// TIA Portal project "g" (V14) (continued)

       REGION Collect-statistics
           // Operating time cnt. (#t_diff will always be zero, if the feature is disabled)
           #devices[#c].operation_time += SEL(G := #devices[#c].in_operation
                                              AND #conf.enable_operation_time_cnt,
                                              IN0 := 0, IN1 := USINT_TO_UDINT(#t_diff));
           // Count number of devices in operation.
           #info.devices_in_operation += BOOL_TO_UINT(#devices[#c].in_operation);
           // Count number of devices in standby.
           #info.devices_standby +=
           BOOL_TO_UINT(#devices[#c].available
                        AND NOT #devices[#c].Q); // NOT #devices[#c].in.in_operation
           // Count number of devices started.
           #info.devices_started += BOOL_TO_UINT(#devices[#c].Q);
       END_REGION
   END_FOR;

   // Some info (for hmi)
   #settings.info.total := DINT_TO_UINT(#upper - #lower + 1);

   // If for some reason, the number operating devies can be limited to less
   // then available
   #settings.max_devices_same_time := // A setting.
   LIMIT(MN := 1,
         IN := #settings.max_devices_same_time,
         MX := #settings.info.total);

   // Force min value for param.
   #settings.max_diff_operating.sec :=
   MAX(IN1 := 60, IN2 := #settings.max_diff_operating.sec);

   // Timers for adding and removing devices for operation.

   #timer_stop.TON(IN := #input < #settings.stop.limit AND NOT #reset_timers,
                   PT := #settings.stop.delay,
                   Q => #timer_stop_q);
   #timer_start.TON(IN := #input > #settings.start.limit AND NOT #reset_timers,
                    PT := #settings.start.delay,
                    Q => #timer_start_q);

   REGION start-stopp
       // Stoping a device
       IF NOT #settings.bypass // The bypass-function turn on all outputs. 
           AND #candidates.stop.index <> #NO_CANDIDATE // A device is available 
           AND (#info.devices_in_operation > 1 // Can't remove last device in operation
           (* *)OR NOT #conf.at_least_one)  // Possible to disable the feature
           AND (
           (* *)#info.devices_in_operation > #settings.max_devices_same_time
           (* *)OR #timer_stop_q // If #input below a certain value for a certain time
           (* *)OR #settings.stop.force  // Used to stop the next device (hmi)
           (* *)OR #boost_start < 0)
       THEN
           #devices[#candidates.stop.index].Q := false; // Disable one device
           RESET_TIMER(#timer_stop);
           #oper := -1;
           // Increase var until zero.
           #boost_start := SEL(G := #boost_start < 0, IN0 := 0, IN1 := #boost_start + 1);

           // Start a devices.
       ELSIF #candidates.start.index <> #NO_CANDIDATE // A device is available 
           AND #info.devices_in_operation < #settings.max_devices_same_time
           AND #input > 0 AND (
           (* *)#info.devices_in_operation < 1 // At least one device operating
           (*      *)AND #conf.at_least_one // Possible to disable the feature
           (* *)OR #timer_start_q // If #input above a certain value for a certain time
           (* *)OR #settings.start.force // Used to starp the next device (hmi)
           (* *)OR #boost_start > 0)
       THEN
           #devices[#candidates.start.index].Q := true; // Enable one more device
           RESET_TIMER(#timer_start);
           #oper := 1;
           // Decrease var until zero.
           #boost_start := SEL(G := #boost_start > 0, IN0 := 0, IN1 := #boost_start - 1);

           // Change operating device, if the operating-time between two devies is to large.
       ELSIF #settings.max_diff_operating.enable
           AND #candidates.start.index <> #NO_CANDIDATE // A candidate is available to be started
           AND #candidates.stop.index <> #NO_CANDIDATE // A candidate is available to be stoped
           AND (#candidates.stop.operation_time - #candidates.start.operation_time >
           (* *)#settings.max_diff_operating.sec) // And the difference is to large.
       THEN
           // Stop the device with most operating time and start the devices with
           // least operating time.
           #devices[#candidates.stop.index].Q := false;
           #devices[#candidates.start.index].Q := true;
       END_IF;
   END_REGION

   // Update vars, after start or stop a device. (above)
   #info.devices_in_operation += SINT_TO_UINT(#oper);
   #info.devices_started += SINT_TO_UINT(#oper);
   #info.devices_standby -= SINT_TO_UINT(#oper);

   // Transfer values to hmi-vars
   #settings.info.in_operation := #info.devices_in_operation;
   #settings.info.started := #info.devices_started;
   #settings.info.standby := #info.devices_standby;

   #settings.info.input := #input;

   // Information has been recived, so now back to default values.
   #set := -1;
   #settings.start.force := false;
   #settings.stop.force := false;
   #settings.boostStart.reset := false;

   // https://github.com/rexhip/
END_FUNCTION_BLOCK

// folder: Library/Alternating/Load balancer/Blocks and UDT's/Internal

FUNCTION "boost_start" : Void   // FC25, SCL
{ S7_Optimized_Access := 'TRUE' }
VERSION : 0.1
   VAR_INPUT
      t_diff : USInt;
      start : Bool;
   END_VAR
   VAR_OUTPUT
      reset_timers : Bool;
   END_VAR
   VAR_IN_OUT
      devices : Array[*] of "load_balancer_device_udt";
      settings : "load_balancer_settings_udt";
      info : "load_balancer_info_udt";
      boost_start : SInt;
      set : SInt;
   END_VAR
   VAR_TEMP
      c : DInt;
      u : DInt;
      lower : DInt;
   END_VAR
BEGIN
   #lower := LOWER_BOUND(ARR := #devices, DIM := 1);
   FOR #c := #lower TO UPPER_BOUND(ARR := #devices, DIM := 1) DO

       #u := #c - #lower + 1; // #u start at 1, increasing by 1 for each iteration.
       IF #settings.boostStart.reset THEN
           // Reset stastic, on how many devices is operating same time.
           #devices[#c].z.n_cnt := 0;
       ELSIF #settings.info.started = #u THEN
           // Log how many devices is operating same time, most fequently.
           #devices[#c].z.n_cnt += #t_diff;
       END_IF;

       // Change how many devices to boost start at startup, based on how many
       // devices is most commenly used.
       IF #settings.boostStart.auto
           AND #devices[#c].z.n_cnt >
           (* *)#devices[#lower + #settings.boostStart.devices - 1].z.n_cnt
       THEN
           #settings.boostStart.devices := DINT_TO_USINT(#u);
       END_IF;
   END_FOR;

   // Set a number of operating devices. (Without waiting for the input and the timers)
   IF #set > -1 THEN
       #boost_start := #set - UINT_TO_SINT(#info.devices_started);

       // Do boost start when input change away from zero.    
   ELSIF #settings.boostStart.enable // HMI enable.
       AND #start
       AND #set = -1
   THEN
       #boost_start :=
       UINT_TO_SINT(#settings.boostStart.devices - #info.devices_started);
   END_IF;
   // #set is put back to -1 at the bottom of the block.

   // MN: Devies started to be stopped.
   // MX: Devices available for start. 
   #boost_start := LIMIT(MN := - UINT_TO_SINT(#info.devices_started),
                         IN := #boost_start,
                         MX := UINT_TO_SINT(#info.devices_standby));

   #reset_timers := #boost_start <> 0 OR #set <> -1; // Reset timers.
END_FUNCTION

// folder: Library/Alternating/Two outputs

FUNCTION_BLOCK "twoOutpus"   // FB23, SCL
{ S7_Optimized_Access := 'TRUE' }
VERSION : 0.1
   VAR_INPUT
      iStartOne : Bool;
      iStartBoth : Bool;
      iavailable1 : Bool := true;
      iavailable2 : Bool := true;
   END_VAR
   VAR_OUTPUT
      q1 : Bool;
      q2 : Bool;
   END_VAR
   VAR RETAIN
      next : SInt := 1;
   END_VAR
   VAR
      ftrig_in : F_TRIG;
   END_VAR
BEGIN
   // Alternating two outputs.

   #ftrig_in(CLK := #iStartOne);

   // Change #next if not available.
   IF NOT #iavailable1 AND #iavailable2 THEN
       #next := 2;
   ELSIF NOT #iavailable2 AND #iavailable1 THEN
       #next := 1;

   // Swap which one to start next time.
   ELSIF #ftrig_in.Q AND NOT #iStartBoth THEN
       #next := SEL(G := #next = 1,
                    IN0 := 1, IN1 := 2);

   // Make sure that value is valid, 1 or 2.    
   ELSIF #next <> 1 AND #next <> 2 THEN
       #next := 1;
   END_IF;

   #q1 := (#next = 1 AND #iStartOne OR #iStartBoth) AND #iavailable1;
   #q2 := (#next = 2 AND #iStartOne OR #iStartBoth) AND #iavailable2;
END_FUNCTION_BLOCK

// folder: Library/Conversion/time and real

FUNCTION "real2time_format" : Time   // FC1, SCL
{ S7_Optimized_Access := 'TRUE' }
VERSION : 0.1
   VAR_INPUT
      in : Real;
      format : SInt;   // 1=ms, 2=sec, 3=min, 4=h, 5=day
   END_VAR
BEGIN
   // PT-max: 24 days, 20 hours, 31 min, 23 sec and 647 ms.

   // Format: 1=ms, 2=sec, 3=min, 4=h, 5=day

   #real2time_format := T#0s;
   CASE #format OF
       1:  // ms
           #real2time_format := T_CONV(REAL_TO_DINT(#in));
       2:  // Sec
           #real2time_format := T_CONV(REAL_TO_DINT(#in * 1000));
       3:  // Min
           #real2time_format := T_CONV(REAL_TO_DINT(#in * 60000)); //  1000*60
       4:  // Hours
           #real2time_format := T_CONV(REAL_TO_DINT(#in * 3600000)); // 1000*60*60
       5:  // Days
           #real2time_format := T_CONV(REAL_TO_DINT(#in * 86400000)); // 1000*60*60*24
   END_CASE;
END_FUNCTION

FUNCTION "time2real_format" : Real   // FC2, SCL
{ S7_Optimized_Access := 'TRUE' }
VERSION : 0.1
   VAR_INPUT
      in : Time;
      format : SInt;   // 1=ms, 2=sec, 3=min, 4=h, 5=day
   END_VAR
BEGIN
   // PT-max: 24 days, 20 hours, 31 min, 23 sec and 647 ms.

   // Format: 1=ms, 2=sec, 3=min, 4=h, 5=day

   #time2real_format := 0;
   CASE #format OF
       1:  // ms
           #time2real_format := DINT_TO_REAL(T_CONV(#in));
       2:  // Sec
           #time2real_format := DINT_TO_REAL(T_CONV(#in)) / 1000;
       3:  // Min
           #time2real_format := DINT_TO_REAL(T_CONV(#in)) / 60000; // 1000*60
       4:  // Hours
           #time2real_format := DINT_TO_REAL(T_CONV(#in)) / 3600000; // 1000*60*60
       5:  // Days
           #time2real_format := DINT_TO_REAL(T_CONV(#in)) / 86400000; // 1000*60*60*24
   END_CASE;
END_FUNCTION

FUNCTION "time_to_real" : Real   // FC28, SCL
{ S7_Optimized_Access := 'TRUE' }
VERSION : 0.1
   VAR_INPUT
      in : Time;
   END_VAR
BEGIN

   #time_to_real := DINT_TO_REAL(T_CONV( #in)) / 1000;
END_FUNCTION

FUNCTION "real_to_time" : Time   // FC29, SCL
{ S7_Optimized_Access := 'TRUE' }
VERSION : 0.1
   VAR_INPUT
      in : Real;
   END_VAR
BEGIN

   #real_to_time := T_CONV(REAL_TO_DINT(#in * 1000));
END_FUNCTION

// folder: Library/Conversion/time_to_str

FUNCTION "tStr" : String   // FC30, SCL
{ S7_Optimized_Access := 'TRUE' }
VERSION : 0.1
   VAR_INPUT
      in : Time;   // Time to be converted in to string.
   END_VAR
   VAR_TEMP
      t : DTL;
      dayOrHour : Bool;
   END_VAR
BEGIN
   // Time to string.

   #t += #in; // Implicit convert to dtl.
   #t.DAY -= 1; 
   #tStr := ''; 

   IF #t.DAY <> 0 THEN
       #tStr := CONCAT(IN1 := RIGHT
                              (IN := S_CONV(#t.DAY),
                               L := 1 + BOOL_TO_INT(#t.DAY > 9)),
                              IN2 := ', ');
   END_IF;
   IF #t.HOUR <> 0 OR LEN(#tStr) <> 0 THEN
       #tStr := CONCAT(IN1 := #tStr,
                              IN2 := RIGHT
                              (IN := S_CONV(#t.HOUR),
                               L := 1 + BOOL_TO_INT(#t.HOUR > 9)),
                              IN3 := ':');
   END_IF;
   #tStr := CONCAT(IN1 := #tStr,
                          IN2 := RIGHT
                          (IN := S_CONV(#t.MINUTE),
                           L := 1 + BOOL_TO_INT(#t.MINUTE > 9)),
                          IN3 := ':');
   #tStr := CONCAT(IN1 := #tStr,
                          IN2 := RIGHT
                          (IN := S_CONV(#t.SECOND),
                           L := 1 + BOOL_TO_INT(#t.SECOND > 9)));

   // https://github.com/rexhip/
END_FUNCTION

// folder: Library/Filters

FUNCTION_BLOCK "digitalRippleFilter"   // FB15, SCL
{ S7_Optimized_Access := 'TRUE' }
VERSION : 0.1
   VAR_INPUT
      in : Bool;
      pt_on : Time;
      pt_off : Time;
   END_VAR
   VAR_OUTPUT
      Q : Bool;
   END_VAR
   VAR
      ton : TON_TIME;
      tof : TOF_TIME;
   END_VAR
BEGIN
   // Filter noice of a digital input signal.

   #ton(IN := #in, PT := #pt_on);

   #tof(IN := #ton.Q OR #tof.Q AND #in,
        PT := #pt_off,
        Q => #Q);
END_FUNCTION_BLOCK

FUNCTION "movingAverageFilter" : Void   // FC7, SCL
{ S7_Optimized_Access := 'TRUE' }
VERSION : 0.1
   VAR_INPUT
      in : Real;
   END_VAR
   VAR_IN_OUT
      filterConst : Real;   // 0=off.
      Q : Real;
   END_VAR
   VAR_TEMP
      z : LReal;
   END_VAR
BEGIN
   // Running average smoothing filter.
   //  - Filter constant has to greater then zero
   //  - PLC scan time will affect the filter.

   IF #filterConst = 0 THEN // Zero -> disable filter 
       #Q := #in;
   ELSE
       #filterConst := MAX(IN1 := 0, IN2 := #filterConst);
       // Creating a number betwwen zero and less then one.
       #z := -1 / REAL_TO_LREAL(#filterConst + 1); 
       #Q := LREAL_TO_REAL(#z * REAL_TO_LREAL(#Q)
                           + (1 - #z) * REAL_TO_LREAL(#in));
   END_IF;
END_FUNCTION

// folder: Library/IO-handeling/Analog in/Blocks

FUNCTION_BLOCK "analogIn_fb"   // FB18, SCL
{ S7_Optimized_Access := 'TRUE' }
VERSION : 0.1
   VAR_INPUT
      in : Int;
   END_VAR
   VAR RETAIN
      aiUdt : "analogInUdt";
   END_VAR
   VAR
      normX : "normXAnalogUdt";
   END_VAR
BEGIN

   "analogIn"(in := #in, aiUdt := #aiUdt, normX := #normX);
END_FUNCTION_BLOCK

FUNCTION "analogIn" : Void   // FC4, SCL
TITLE = Analog input
{ S7_Optimized_Access := 'TRUE' }
VERSION : 0.1
   VAR_INPUT
      in : Int;
   END_VAR
   VAR_IN_OUT
      aiUdt : "analogInUdt";
      normX : "normXAnalogUdt";
   END_VAR
   VAR_TEMP
      u : Real;
      x : Real;
      y : Real;
      "e" : Int;
   END_VAR
BEGIN
   // Analog input scaling.

   #u := NORM_X(MIN := #normX.rawMin, VALUE := #in, MAX := #normX.rawMax);
   "movingAverageFilter"(in := #u,
                         filterConst := #aiUdt.filterConst,
                         Q := #aiUdt.unitInterval);
   IF #aiUdt.sim THEN
       ; // A simulated value can be set directly to #aiUdt.Q and #aiUdt.Error
   ELSE
       // Scale back up to raw-value to check if outside error limits.
       #x := SCALE_X(MIN := #normX.rawMin, MAX := #normX.rawMax,
                     VALUE := #aiUdt.unitInterval);
       #aiUdt.Error := #x < #normX.errorLimMin OR #x > #normX.errorLimMax;
       // Log the time when the error occurred.
       IF #aiUdt.Error AND NOT #aiUdt.zOldError THEN
           #"e" := RD_LOC_T(#aiUdt.ErrorTime);
       END_IF;

       IF #aiUdt.Error THEN
           #y := SINT_TO_REAL(#aiUdt.errorAction) / 100;
       ELSIF #aiUdt.forceInsideScale THEN
           #y := LIMIT(MN := 0, IN := #aiUdt.unitInterval, MX := 1);
       ELSE
           #y := #aiUdt.unitInterval;
       END_IF;
       #aiUdt.Q := SCALE_X(MIN := #aiUdt.scaleMin, MAX := #aiUdt.scaleMax,
                           VALUE := #y ) * #aiUdt.gain + #aiUdt.offset;
   END_IF;
   #aiUdt.zOldError := #aiUdt.Error;

   // ( https://github.com/rexhip/ )
END_FUNCTION

FUNCTION "analogInAndAlarms" : Void   // FC6, SCL
{ S7_Optimized_Access := 'TRUE' }
VERSION : 0.1
   VAR_INPUT
      in : Int;
   END_VAR
   VAR_IN_OUT
      aiUdt : "analogInAndAlarmsUdt";
      ioGlobal : "ioGlobal_FB";
   END_VAR
   VAR CONSTANT
      VALUE_LESS_THEN_LIM : SInt := 1;
      VALUE_GREATER_THEN_LIM : SInt := 2;
   END_VAR
BEGIN
   // Analog input with alarm handling. 

   REGION Input handling
       // A id for each io
       #ioGlobal.z.ioIdCnt += 1;

       // Disable all simulations.
       #aiUdt.ai.sim := #aiUdt.ai.sim AND NOT #ioGlobal.info2ioBlocks.disableAllSim;

       IF #aiUdt.execAiLogic THEN // Execute analog input logic
           "analogIn"(in := #in,
                      aiUdt := #aiUdt.ai,
                      normX := #ioGlobal.normX);
       END_IF;
       // Count number of errors
       #ioGlobal.collectInfo.errorCnt += BOOL_TO_UINT(#aiUdt.ai.Error);;
       // Count active simulations 
       #ioGlobal.collectInfo.activeSimCnt += BOOL_TO_UINT(#aiUdt.ai.sim);
   END_REGION

   REGION Alarms  
   // Connecting ioGlobal functions with each alarm.
   "ioGlobalAlarmLinking"(alarm := #aiUdt.alarmHH, ioGlobal := #ioGlobal);
   "ioGlobalAlarmLinking"(alarm := #aiUdt.alarmH, ioGlobal := #ioGlobal);
   "ioGlobalAlarmLinking"(alarm := #aiUdt.alarmLL, ioGlobal := #ioGlobal);
   "ioGlobalAlarmLinking"(alarm := #aiUdt.alarmL, ioGlobal := #ioGlobal);

   "alarmReal"(value := #aiUdt.ai.Q, // HH alarm
               action := #VALUE_GREATER_THEN_LIM,
               disable := false,
               runtimeDiff := #ioGlobal.info2ioBlocks.runtimeDiff,
               alarm := #aiUdt.alarmHH);
   "alarmReal"(value := #aiUdt.ai.Q,// H alarm
               action := #VALUE_GREATER_THEN_LIM,
               disable := #aiUdt.alarmHH.Q,
               runtimeDiff := #ioGlobal.info2ioBlocks.runtimeDiff,
               alarm := #aiUdt.alarmH);
   "alarmReal"(value := #aiUdt.ai.Q, // LL alarm
               action := #VALUE_LESS_THEN_LIM,
               disable := false,
               runtimeDiff := #ioGlobal.info2ioBlocks.runtimeDiff,
               alarm := #aiUdt.alarmLL);
   "alarmReal"(value := #aiUdt.ai.Q, // L alarm
               action := #VALUE_LESS_THEN_LIM,
               disable := #aiUdt.alarmLL.Q,
               runtimeDiff := #ioGlobal.info2ioBlocks.runtimeDiff,
               alarm := #aiUdt.alarmL);
   END_REGION

   REGION HMI-features
       // Copy paste all settings. (HMI)
       IF #aiUdt.hmi.copyAllSettings THEN
           #ioGlobal.copyPaste := #aiUdt;
           #aiUdt.hmi.copyAllSettings := false;
       ELSIF #aiUdt.hmi.pasteAllSettings THEN
           "pasteAnalogInSetting"(src := #ioGlobal.copyPaste, dest := #aiUdt);
           #aiUdt.hmi.pasteAllSettings := false;
       END_IF;

       #aiUdt.hmi.showTag := #ioGlobal.hmi.hmiShowTags;
   END_REGION

   // ( https://github.com/rexhip/ )
END_FUNCTION

FUNCTION "analogInSimple" : Real   // FC13, SCL
{ S7_Optimized_Access := 'TRUE' }
VERSION : 0.1
   VAR_INPUT
      mn : Real;
      in : Int;
      mx : Real;
   END_VAR
   VAR_TEMP
      x : Real;
   END_VAR
BEGIN
   // Analog in 

   #x := NORM_X(MIN := 0, VALUE := #in, MAX := 27648);
   #x := LIMIT(MN := 0, IN := #x, MX := 1);
   #analogInSimple := SCALE_X(MIN := #mn, VALUE := #x, MAX := #mx);

   // ( https://github.com/rexhip/ )
END_FUNCTION

FUNCTION "analogInError" : Bool   // FC14, SCL
{ S7_Optimized_Access := 'TRUE' }
VERSION : 0.1
   VAR_INPUT
      in : Int;
   END_VAR
   VAR_TEMP
      t : Real;
   END_VAR
BEGIN
   // Analog in error (outside limits.)
   #analogInError := #in < -4864 OR #in > 32512;;
END_FUNCTION

FUNCTION "analogInReal" : Void   // FC34, SCL
{ S7_Optimized_Access := 'TRUE' }
VERSION : 0.1
   VAR_INPUT
      in : Real;
      error : Bool;
   END_VAR
   VAR_IN_OUT
      aiUdt : "analogInAndAlarmsUdt";
      ioGlobal : "ioGlobal_FB";
   END_VAR
   VAR_TEMP
      dommy : Int;
      u : Real;
   END_VAR
BEGIN
   // Analog input 
   // Wrapper to use analog input block with real input.
   // 
   #aiUdt.ai.Error := #error;

   IF #aiUdt.ai.sim THEN
       ; // A simultated value may be set directly at: #ai.ai.Q
   ELSE
       #u := #in * #aiUdt.ai.gain + #aiUdt.ai.offset;
       "movingAverageFilter"(in := #u,
                             filterConst := #aiUdt.ai.filterConst,
                             Q := #aiUdt.ai.Q);
   END_IF;

   #aiUdt.execAiLogic := false;
   "analogInAndAlarms"(in := #dommy,
                       aiUdt := #aiUdt,
                       ioGlobal := #ioGlobal);

   // ( https://github.com/rexhip/ )
END_FUNCTION

// folder: Library/IO-handeling/Analog in/internal

FUNCTION "ioGlobalAlarmLinking" : Void   // FC3, SCL
{ S7_Optimized_Access := 'TRUE' }
VERSION : 0.1
   VAR_IN_OUT
      alarm : "alarmRealUdt";
      ioGlobal : "ioGlobal_FB";
   END_VAR
BEGIN
   // Connecting ioGlobal functions with valueAlarm.

   // Acknowle alarm
   #alarm.ack := #ioGlobal.info2ioBlocks.ackAllAlarms;

   // Count active alarms
   #ioGlobal.collectInfo.activeAlarmsCnt += BOOL_TO_UINT(#alarm.Q);
   // Count unacknowledged alarms
   #ioGlobal.collectInfo.unacknowledgedAlarmsCnt +=
   BOOL_TO_UINT(#alarm.Q AND NOT #alarm.memAck);

   // ( https://github.com/rexhip/ )
END_FUNCTION

FUNCTION "pasteAnalogInSetting" : Void   // FC20, SCL
{ S7_Optimized_Access := 'TRUE' }
VERSION : 0.1
   VAR_IN_OUT
      src : "analogInAndAlarmsUdt";
      dest : "analogInAndAlarmsUdt";
   END_VAR
BEGIN
   // Select only the settings and not values from the 
   // udt's and transfer them from src to dest.

   #dest.ai.offset := #src.ai.offset ;
   #dest.ai.errorAction := #src.ai.errorAction ;
   #dest.ai.gain := #src.ai.gain ;
   #dest.ai.filterConst := #src.ai.filterConst ;
   #dest.ai.forceInsideScale := #src.ai.forceInsideScale ;
   #dest.ai.scaleMax := #src.ai.scaleMax ;
   #dest.ai.scaleMin := #src.ai.scaleMin ;

   "pasteAlarmSetting"(src := #src.alarmHH, dest := #dest.alarmHH);
   "pasteAlarmSetting"(src := #src.alarmH,  dest := #dest.alarmH);
   "pasteAlarmSetting"(src := #src.alarmLL, dest := #dest.alarmLL);
   "pasteAlarmSetting"(src := #src.alarmL,  dest := #dest.alarmL);
END_FUNCTION

FUNCTION "pasteAlarmSetting" : Void   // FC21, SCL
{ S7_Optimized_Access := 'TRUE' }
VERSION : 0.1
   VAR_IN_OUT
      src : "alarmRealUdt";
      dest : "alarmRealUdt";
   END_VAR
BEGIN

   #dest.enable := #src.enable;
   #dest.autoAck := #src.autoAck ;
   #dest.delay := #src.delay ;
   #dest.hyst := #src.hyst ;
   #dest.lim := #src.lim ;
END_FUNCTION

// folder: Library/IO-handeling/Analog out

FUNCTION "analogOut" : Void   // FC9, SCL
{ S7_Optimized_Access := 'TRUE' }
VERSION : 0.1
   VAR_OUTPUT
      q : Int;
   END_VAR
   VAR_IN_OUT
      aoUdt : "analogOutUdt_1";
      ioGlobal : "ioGlobal_FB";
   END_VAR
   VAR_TEMP
      x : Real;
      y : Real;
   END_VAR
BEGIN
   // Analog out 

   // - failSafe: Output will go to a predefined value set by
   //   failSafeValue (%), this can be used for emergency stop.
   //   Simulation will not work when failSafe is activated.

   // A id for each io
   #ioGlobal.z.ioIdCnt += 1;

   IF #ioGlobal.info2ioBlocks.disableAllSim THEN
       #aoUdt.simEnable := false;
   END_IF;

   IF #aoUdt.failSafe THEN
       #x := SINT_TO_REAL(#aoUdt.failSafeValue) / 100 ; // [%]
   ELSE
       IF #aoUdt.simEnable THEN
           #y := #aoUdt.simValue;
       ELSIF #aoUdt.interlook THEN
           #y := 0;
       ELSE
           #y := #aoUdt.in;
       END_IF;
       #x := NORM_X(MIN := #aoUdt.scaleMin, VALUE := #y,
                    MAX := #aoUdt.scaleMax);
       #aoUdt.simValue := #y;
   END_IF;
   #x := LIMIT(MN := 0, IN := #x, MX := 1);
   #q := SCALE_X(MIN := #ioGlobal.normX.rawMin, VALUE := #x,
                     MAX := #ioGlobal.normX.rawMax);

   #ioGlobal.collectInfo.activeSimCnt += BOOL_TO_UINT(#aoUdt.simEnable);

   // ( https://github.com/rexhip/ )
END_FUNCTION

FUNCTION "analogOutSimple" : Int   // FC22, SCL
{ S7_Optimized_Access := 'TRUE' }
VERSION : 0.1
   VAR_INPUT
      in : Real;   // Percent
   END_VAR
   VAR_TEMP
      x : Real;
   END_VAR
BEGIN
   // Simple analog unipolar output

   // Input:  per cent.
   // Output: Siemens unipolar scale.

   #x := LIMIT(MN := 0, IN := #in / 100, MX := 1);
   #analogOutSimple := SCALE_X(MIN := 0, VALUE := #x, MAX := 27648);

   // ( https://github.com/rexhip/ )
END_FUNCTION

// folder: Library/IO-handeling/Common functions

FUNCTION_BLOCK "ioGlobal_FB"   // FB7, SCL
{ S7_Optimized_Access := 'TRUE' }
VERSION : 0.1
   VAR
      hmi : "ioGlobalUdt";
      z_internal_timer : IEC_TIMER;
      z_internal : Struct
         fs : Bool := TRUE;
         timer_mem : Time;
      END_STRUCT;
      collectInfo : Struct
         activeSimCnt : UInt;
         activeAlarmsCnt : UInt;
         unacknowledgedAlarmsCnt : UInt;
         errorCnt : UInt;
      END_STRUCT;
      info2ioBlocks : Struct
         runtimeDiff : Time;
         ackAllAlarms : Bool;
         disableAllSim : Bool;
         firstScan : Bool := TRUE;
      END_STRUCT;
      z : Struct
         ioIdCnt : UInt;
      END_STRUCT;
      copyPaste : "analogInAndAlarmsUdt";
      normX : "normXAnalogUdt";
   END_VAR
BEGIN
   // ioGlobal: This block handels common function for io, eg:
   //  - Count active simulations
   //  - Disable all simulations
   //  - Count active alarms
   //  - Ack. all active alarms

   // Calculate time of each plc scan.
   #z_internal_timer.TON(IN := NOT #z_internal_timer.Q, PT := T#24d);
   IF #z_internal_timer.ET <> #z_internal.timer_mem THEN
       #info2ioBlocks.runtimeDiff := #z_internal_timer.ET - #z_internal.timer_mem;
   END_IF;
   #z_internal.timer_mem := #z_internal_timer.ET;

   // First scan
   #info2ioBlocks.firstScan := #z_internal.fs;
   #z_internal.fs := false;

   // Common information to all io-blocks.
   #info2ioBlocks.ackAllAlarms := #hmi.ackAllAlarms;
   #info2ioBlocks.disableAllSim := #hmi.disableAllSim;
   // Make sure that ack only happens once.
   #hmi.ackAllAlarms := false;
   #hmi.disableAllSim := false;

   // Information from io-blocks.
   #hmi.totalActiveAlarms := #collectInfo.activeAlarmsCnt;
   #hmi.totalActiveSim := #collectInfo.activeSimCnt;
   #hmi.totalUnacknowledgedAlarms := #collectInfo.unacknowledgedAlarmsCnt;
   #hmi.totalErrors := #collectInfo.errorCnt;
   // Reset the counter for new collection of info on next scan.
   #collectInfo.activeAlarmsCnt := 0;
   #collectInfo.activeSimCnt := 0;
   #collectInfo.unacknowledgedAlarmsCnt := 0;
   #collectInfo.errorCnt := 0;

   // ioId io-id
   #z.ioIdCnt := 0;

   // ( https://github.com/rexhip/ )
END_FUNCTION_BLOCK

FUNCTION "alarmBoolSimple" : Void   // FC5, SCL
{ S7_Optimized_Access := 'TRUE' }
VERSION : 0.1
   VAR_INPUT
      in : Bool;
   END_VAR
   VAR_IN_OUT
      alarm : "alarmBoolSimpleUdt";
   END_VAR
BEGIN
   // Simple digital alarm 

   IF #alarm.enable THEN
       IF #alarm.Q THEN
           #alarm.memAck := #alarm.memAck OR #alarm.ack; // Acknowledge
           IF NOT #alarm.in AND (
               #alarm.autoAck
               OR #alarm.memAck AND NOT #alarm.dobleAck
               OR #alarm.ack AND #alarm.dobleAck)
           THEN
               #alarm.Q := false;
           END_IF;
       ELSIF #alarm.in THEN
           #alarm.Q := true;
           #alarm.memAck := false;
       END_IF;
       #alarm.ack := false;

   ELSE // Alarm is disabled
       #alarm.Q := false;
   END_IF;
END_FUNCTION

FUNCTION "alarmReal" : Void   // FC11, SCL
{ S7_Optimized_Access := 'TRUE' }
VERSION : 0.1
   VAR_INPUT
      value : Real;   // Value that will be compared
      action : SInt;   // 1=Greater then, 2=less then
      disable : Bool;   // diable alarm
   END_VAR
   VAR_IN_OUT
      runtimeDiff : Time;   // Time of last program scan, used for internal timer
      alarm : "alarmRealUdt";
   END_VAR
   VAR_TEMP
      tmpQset : Bool;
      tmpQrst : Bool;
   END_VAR
   VAR CONSTANT
      LESS_THEN : SInt := 1;
      GREATER_THEN : SInt := 2;
   END_VAR
BEGIN
   // Value alarm

   #alarm.value := #value;
   #alarm.action := #action;

   IF #alarm.enable AND NOT #disable THEN
       CASE #action OF
           #LESS_THEN: // (1)
               #tmpQset := #value < #alarm.lim;
               #tmpQrst := #value > #alarm.lim + #alarm.hyst;
           #GREATER_THEN: // (2)
               #tmpQset := #value > #alarm.lim;
               #tmpQrst := #value < #alarm.lim - #alarm.hyst;
       END_CASE;
       IF #alarm.Q THEN  // if alarm has been activated.
           #alarm.memAck := #alarm.memAck OR #alarm.ack; // Acknowledge
           IF #tmpQrst AND (
               #alarm.autoAck
               OR #alarm.memAck AND NOT #alarm.dobleAck
               OR #alarm.ack AND #alarm.dobleAck)
           THEN
               #alarm.Q := false;
           END_IF;
       ELSE  // Not #alarm.Q
           IF #tmpQset THEN
               #alarm.delayEt += #runtimeDiff;
               IF #alarm.delayEt >= #alarm.delay THEN
                   #alarm.Q := true;
                   #alarm.memAck := false;
               END_IF;
           ELSE
               #alarm.delayEt := T#0s;
           END_IF;
       END_IF;
       #alarm.ack := false;

   ELSE // Alarm disabled
       #alarm.Q := false;
       #alarm.delayEt := T#0s;
   END_IF;

   // ( https://github.com/rexhip/ )
END_FUNCTION

FUNCTION "setUnipolar" : Void   // FC18, SCL
{ S7_Optimized_Access := 'TRUE' }
VERSION : 0.1
   VAR_IN_OUT
      unipolar : "normXAnalogUdt";
   END_VAR
BEGIN
   // Set values for analog input and output to
   // unipolar.

   #unipolar.rawMin := 0;
   #unipolar.rawMax := 27648;

   // Outside limits bellow will generate error.
   #unipolar.errorLimMin := -4864;
   #unipolar.errorLimMax := 32512;
END_FUNCTION

FUNCTION "setAnalogType" : "normXAnalogUdt"   // FC19, SCL
{ S7_Optimized_Access := 'TRUE' }
VERSION : 0.1
   VAR_INPUT
      select : Int;
   END_VAR
   VAR_TEMP
      dommy : "normXAnalogUdt";
   END_VAR
BEGIN
   // Set values for analog input and output 

   CASE #select OF
       1:  // Siemens unipolar
           #setAnalogType.rawMin := 0;
           #setAnalogType.rawMax := 27648;
           #setAnalogType.errorLimMin := -4864;
           #setAnalogType.errorLimMax := 32512;
       2:  // Siemens bipolar
           #setAnalogType.rawMin := -27648;
           #setAnalogType.rawMax := 27648;
           #setAnalogType.errorLimMin := -32512;
           #setAnalogType.errorLimMax := 32512;
       3:  // Wago - 750-496  - 0/4-20 mA
           #setAnalogType.rawMin := 0;
           #setAnalogType.rawMax := 30832;
           #setAnalogType.errorLimMin := -773;
           #setAnalogType.errorLimMax := 32763;
           // 4:  
           //  #setAnalogType.min := ;
           //  #setAnalogType.max := ;
           //  #setAnalogType.errorLimMin := ;
           //  #setAnalogType.errorLimMax := ;
       ELSE
           #setAnalogType := #dommy;
   END_CASE;
END_FUNCTION

// folder: Library/IO-handeling/Common functions/z Dev

FUNCTION "syncAlarmReal" : Void   // FC26, SCL
{ S7_Optimized_Access := 'TRUE' }
VERSION : 0.1
   VAR_IN_OUT
      prim : "alarmRealUdt";
      sec : "alarmRealUdt";
      memory : "alarmRealUdt";
   END_VAR
BEGIN

   #prim.value := #sec.value;
   #prim.action := #sec.action;

   "syncReal"(prim := #prim.lim ,
              sec := #sec.lim ,
              memory := #memory.lim);

   "syncBool"(prim := #prim.Q,
              sec := #sec.Q,
              memory := #memory.Q);
END_FUNCTION

// folder: Library/IO-handeling/Digital in

FUNCTION "digitalIn" : Void   // FC10, SCL
{ S7_Optimized_Access := 'TRUE' }
VERSION : 0.1
   VAR_INPUT
      in : Bool;
   END_VAR
   VAR_IN_OUT
      diUdt : "digitalInUdt";
      ioGlobal : "ioGlobal_FB";
   END_VAR
   VAR_TEMP
      "e" : Int;
      tmpQ : Bool;
      tmpIn : Bool;
   END_VAR
BEGIN
   // Digital input ( https://github.com/rexhip/ )

   // A id for each io
   #ioGlobal.z.ioIdCnt += 1;

   IF #diUdt.sim THEN
       #diUdt.delayEt := T#0ms;
   ELSE
       #tmpQ := #diUdt.Q;
       #tmpIn := #in XOR #diUdt.invert;
       IF #tmpIn AND NOT #diUdt.Q THEN
           #diUdt.delayEt += #ioGlobal.info2ioBlocks.runtimeDiff;
       ELSIF NOT #tmpIn THEN
           #diUdt.delayEt := T#0ms;
       END_IF;
       #diUdt.Q := #diUdt.delayEt >= #diUdt.delay;

       // Logging - the time the input change state.
       IF #diUdt.Q AND NOT #tmpQ THEN
           #"e" := RD_LOC_T(#diUdt.timeOn);
       ELSIF NOT #diUdt.Q AND #tmpQ THEN
           #"e" := RD_LOC_T(#diUdt.timeOff);
       END_IF;
   END_IF;

   "alarmBoolSimple"(in := #diUdt.Q, alarm := #diUdt.alarm);

   // Count alarms, errors and simulations.
   #ioGlobal.collectInfo.activeAlarmsCnt += BOOL_TO_UINT(#diUdt.alarm.Q);
   #ioGlobal.collectInfo.errorCnt += BOOL_TO_UINT(#diUdt.Error);;
   #ioGlobal.collectInfo.activeSimCnt += BOOL_TO_UINT(#diUdt.sim);

   // ( https://github.com/rexhip/ )
END_FUNCTION

// folder: Library/IO-handeling/Digital out

FUNCTION "digitalOut" : Void   // FC8, SCL
{ S7_Optimized_Access := 'TRUE' }
VERSION : 0.1
   VAR_OUTPUT
      Out : Bool;
   END_VAR
   VAR_IN_OUT
      doUdt : "digitalOutUdt";
      ioGlobal : "ioGlobal_FB";
   END_VAR
   VAR_TEMP
      t : Bool;
   END_VAR
BEGIN
   // Digital out
   //
   // - For most application a analog output block is not needed. However
   //
   // - failSafe: Output will go to a predefined value set by failSafeValue (%),
   //   this can be used for emergency stop, simulation will not work when
   //   failSafe is activated.

   // A id for each io
   #ioGlobal.z.ioIdCnt += 1;

   IF #doUdt.disableSim OR #ioGlobal.info2ioBlocks.disableAllSim THEN
       #doUdt.simEnable := false;
   END_IF;

   IF #doUdt.failSafe THEN
       #t := #doUdt.failSafeValue;
   ELSE
       #t := SEL(G := #doUdt.simEnable,
                 IN0 := #doUdt.in XOR #doUdt.invert,
                 IN1 := #doUdt.simValue);
   END_IF;
   #doUdt.simValue := #Out := #t;

   #ioGlobal.collectInfo.activeSimCnt += BOOL_TO_USINT(#doUdt.simEnable);

   // ( https://github.com/rexhip/ )
END_FUNCTION

// folder: Library/IO-handeling/_examples

FUNCTION_BLOCK "_example_analogOutpus"   // FB2, SCL
{ S7_Optimized_Access := 'TRUE' }
VERSION : 0.1
   VAR_OUTPUT
      ao_FV01 : Int;
      ao_FV02 : Int;
      ao_FV03 : Int;
   END_VAR
   VAR_IN_OUT
      ioGlobal : "ioGlobal_FB";
   END_VAR
   VAR RETAIN
      FV01 : "analogOutUdt_1";
      FV02 : "analogOutUdt_1";
   END_VAR
   VAR
      FV03 : Real;
   END_VAR
BEGIN


   "analogOut"(aoUdt := #FV01,
               ioGlobal := #ioGlobal,
               q => #ao_FV01);

   "analogOut"(aoUdt := #FV02,
               ioGlobal := #ioGlobal,
               q => #ao_FV02);

   // Very simple analog output.
   #ao_FV03 := "analogOutSimple"(#FV03);
END_FUNCTION_BLOCK

FUNCTION_BLOCK "_example_digitalOutpus"   // FB4, SCL
{ S7_Optimized_Access := 'TRUE' }
VERSION : 0.1
   VAR_OUTPUT
      do_PX01 : Bool;
      do_PX02 : Bool;
   END_VAR
   VAR_IN_OUT
      ioGlobal : "ioGlobal_FB";
   END_VAR
   VAR RETAIN
      PX01 : "digitalOutUdt";
      PX02 : "digitalOutUdt";
   END_VAR
BEGIN

   "digitalOut"(Out => #do_PX01,
                doUdt := #PX01,
                ioGlobal := #ioGlobal);

   "digitalOut"(Out => #do_PX02,
                doUdt := #PX02,
                ioGlobal := #ioGlobal);
END_FUNCTION_BLOCK

FUNCTION_BLOCK "_example_analogInputs"   // FB5, SCL
{ S7_Optimized_Access := 'TRUE' }
VERSION : 0.1
   VAR_INPUT
      ai_FT12 : Int;
      ai_TT27 : Int;
      value_from_other_source : Real;
   END_VAR
   VAR_IN_OUT
      ioGlobal : "ioGlobal_FB";
   END_VAR
   VAR RETAIN
      FT12 : "analogInAndAlarmsUdt";
      TT27 : "analogInAndAlarmsUdt";
      PT44 : "analogInAndAlarmsUdt";
   END_VAR
BEGIN
   // Analog inputs example. ( https://github.com/rexhip/ )

   // In a real world example the input on this block
   // would be PLC-tags connected to fysical IO.

   "analogInAndAlarms"(in := #ai_FT12,
                       aiUdt := #FT12,
                       ioGlobal := #ioGlobal);
   "analogInAndAlarms"(in := #ai_TT27,
                       aiUdt := #TT27,
                       ioGlobal := #ioGlobal);

   // Value arriving from other source, eg. profinet.
   "analogInReal"(in := #value_from_other_source,
                  error := false, // Should be provided in case comm. error.
                  aiUdt := #PT44,
                  ioGlobal := #ioGlobal);
END_FUNCTION_BLOCK

FUNCTION_BLOCK "_example_digitalInputs"   // FB16, SCL
{ S7_Optimized_Access := 'TRUE' }
VERSION : 0.1
   VAR_INPUT
      di_PAH01 : Bool;
      di_PAH02 : Bool;
   END_VAR
   VAR_IN_OUT
      ioGlobal : "ioGlobal_FB";
   END_VAR
   VAR RETAIN
      PAH01 : "digitalInUdt";
      PAH02 : "digitalInUdt";
   END_VAR
BEGIN

   "digitalIn"(in := #di_PAH01,
               diUdt := #PAH01,
               ioGlobal := #ioGlobal);
   "digitalIn"(in := #di_PAH02,
               diUdt := #PAH02,
               ioGlobal := #ioGlobal);
END_FUNCTION_BLOCK

// folder: Library/Misc/Set reset

FUNCTION "setReset_rd" : Void   // FC15, SCL
{ S7_Optimized_Access := 'TRUE' }
VERSION : 0.1
   VAR_INPUT
      s : Bool;
      r : Bool;
   END_VAR
   VAR_IN_OUT
      q : Bool;
   END_VAR
BEGIN
   // Set-reset (sd = reset dominant)

   IF #r THEN
       #q := false;
   ELSIF #s THEN
       #q := true;
   END_IF;
END_FUNCTION

FUNCTION "setReset_sd" : Void   // FC16, SCL
{ S7_Optimized_Access := 'TRUE' }
VERSION : 0.1
   VAR_INPUT
      s : Bool;
      r : Bool;
   END_VAR
   VAR_IN_OUT
      q : Bool;
   END_VAR
BEGIN
   // Set-reset (sd = reset dominant)

   IF #s THEN
       #q := true;
   ELSIF #r THEN
       #q := false;
   END_IF;
END_FUNCTION

// folder: Library/Misc/operating time

FUNCTION "operatingTime" : Void   // FC12, SCL
{ S7_Optimized_Access := 'TRUE' }
VERSION : 0.1
   VAR_INPUT
      in : Bool;
   END_VAR
   VAR_IN_OUT
      opr : "operatingTimeUdt";
   END_VAR
   VAR_TEMP
      "e" : Int;
      rdSysT : DTL;
   END_VAR
BEGIN
   // This function shouldn't be used with periodical interupts that has longer
   // cycles then 50 secounds.

   // Operating time.
   // (Max value: 2^32 / (24 * 60*60 * 365) = 136 => 136 years.)
   #"e" := RD_SYS_T(#rdSysT);
   #opr.operatingTime +=
   SEL(G := #in, IN0 := 0, IN1 := (#rdSysT.SECOND - #opr.oldSec + 60) MOD 60);
   #opr.oldSec := #rdSysT.SECOND;

   // Start cnt.
   #opr.startCnt += BOOL_TO_UDINT(#in AND NOT #opr.oldIn);
   #opr.oldIn := #in;
END_FUNCTION

// folder: Library/Misc/sync

FUNCTION "syncReal" : Void   // FC17, SCL
{ S7_Optimized_Access := 'TRUE' }
VERSION : 0.1
   VAR_IN_OUT
      prim : Real;   // primary
      sec : Real;   // secoundary
      memory : Real;
   END_VAR
BEGIN
   // Make two variables have the same value. If one change, the
   // value will be transfer to the other one.

   IF #prim = #memory THEN
       #prim := #sec;
   ELSE
       #sec := #prim;
   END_IF;

   #memory := #sec;
END_FUNCTION

FUNCTION "syncBool" : Void   // FC27, SCL
{ S7_Optimized_Access := 'TRUE' }
VERSION : 0.1
   VAR_IN_OUT
      prim : Bool;   // primary
      sec : Bool;   // secoundary
      memory : Bool;
   END_VAR
BEGIN
   // Make two variables have the same value. If one change, the
   // value will be transfer to the other one.

   IF #prim = #memory THEN
       #prim := #sec;
   ELSE
       #sec := #prim;
   END_IF;

   #memory := #sec;
END_FUNCTION

// folder: Library/PID

FUNCTION_BLOCK "pid"   // FB19, SCL
{ S7_Optimized_Access := 'TRUE' }
VERSION : 0.1
   VAR
      pidUdt : "pidUdt";
      pidCompact : PID_Compact;
      oldSec : USInt;
   END_VAR
   VAR_TEMP
      T : DTL;
      "e" : Int;
   END_VAR
BEGIN

   //#e := RD_SYS_T(#T);
   //IF #T.SECOND <> #oldSec THEN
   #pidCompact.Retain.CtrlParams := #pidUdt.pidParam;
   #pidCompact(Setpoint := #pidUdt.sp,
               Input := #pidUdt.pv,
               ManualEnable := #pidUdt.man,
               Output => #pidUdt.mv,
               Error => #pidUdt.error);
   //END_IF;
   //#oldSec := #T.SECOND;
END_FUNCTION_BLOCK

// folder: Library/State machine

FUNCTION_BLOCK "example_stateMachine"   // FB21, SCL
{ S7_Optimized_Access := 'TRUE' }
VERSION : 0.1
   VAR
      state : Int;
      old_state : Int;
      timer1 : TON_TIME;
      timer2 : TON_TIME;
      __condition_1__ : Bool := TRUE;
      __condition_2__ : Bool := TRUE;
      HMI_status : String[100];
   END_VAR
BEGIN
   // State machine with timer example. (https://github.com/rexhip/)

   CASE #state OF
       0:  // Next state after 14 sec. Note that the timer is only one line of code.
           #state += BOOL_TO_INT("timer"(pt := T#14s, t := #timer1));

           #HMI_status := CONCAT(IN1 := 'State 0, remaining time: ',
                                 IN2 := "tStr"("rt"(#timer1)), IN3 := '.');

       1:  // Next state after 7 sec, and '__condition_1__' is true.
           #timer1(IN := true, PT := T#7s);
           #state += BOOL_TO_INT(#timer1.Q AND #__condition_1__);

           // Back to stae 0 if:
           IF "timer"(pt := T#1m50s, t := #timer2) THEN
               #state := 0;
           END_IF;

           #HMI_status := CONCAT(IN1 := 'State 1, Timer1 ', IN2 := "tStr"("rt"(#timer1)),
                                 IN3 := ', Timer2 ', IN4 := "tStr"("rt"(#timer2)));

       2:  // Back to state 0, when '__condition_2__' has been true for 8 sec continuously.
           #timer1(IN := #__condition_2__, PT := T#8s);
           #state := SEL(G := #timer1.Q, IN0 := #state, IN1 := 0);

           #HMI_status := 'State 2.';
   END_CASE;

   IF #state <> #old_state THEN
       RESET_TIMER(#timer1);
       RESET_TIMER(#timer2);
   END_IF;
   #old_state := #state;
END_FUNCTION_BLOCK

FUNCTION "timer" : Bool   // FC23, SCL
{ S7_Optimized_Access := 'TRUE' }
VERSION : 0.1
   VAR_INPUT
      pt : Time;
   END_VAR
   VAR_IN_OUT
      t : TON_TIME;
   END_VAR
BEGIN
   #t(IN := true, PT := #pt);
   #"timer" := #t.Q;
END_FUNCTION

FUNCTION "rt" : Time   // FC31, SCL
{ S7_Optimized_Access := 'TRUE' }
VERSION : 0.1
   VAR_IN_OUT
      "timer" : TON_TIME;
   END_VAR
BEGIN
   // Remaining time
   #rt := #"timer".PT - #"timer".ET;
END_FUNCTION

// folder: Library/Timers

FUNCTION_BLOCK "setResetTimer"   // FB17, SCL
{ S7_Optimized_Access := 'TRUE' }
VERSION : 0.1
   VAR_INPUT
      in : Bool;
      pt : Time;
      set : Bool;
      reset : Bool;
   END_VAR
   VAR_OUTPUT
      q : Bool;
   END_VAR
   VAR
      "timer" : IEC_TIMER;
      timer_q : Bool;
   END_VAR
BEGIN
   // Once the timer has elapsed, the output
   // will stay true until it's reset.

   #"timer".TON(IN := #in, PT := #pt, Q => #timer_q);

   IF #set THEN
       #q := true;
   ELSIF #reset THEN
       #q := false;
   ELSIF #timer_q THEN
       #q := true;
   END_IF;
END_FUNCTION_BLOCK

// folder: Library/Timers/Interval

FUNCTION_BLOCK "Interval"   // FB22, SCL
{ S7_Optimized_Access := 'TRUE' }
VERSION : 0.1
   VAR_INPUT
      in : Bool;   // Activate interval timer
   END_VAR
   VAR_OUTPUT
      Q : Bool;   // Output
      RT : Time;   // Remaining time
   END_VAR
   VAR_IN_OUT
      udt : "intervalUdt";
   END_VAR
   VAR
      N : UDInt;   // Number of cycles
      "timer" : IEC_TIMER;
   END_VAR
   VAR_TEMP
      r : Real;
      t : Time;
      "b" : Bool;
   END_VAR
   VAR CONSTANT
      SECOUNDS : SInt := 1;
   END_VAR
BEGIN
   // When #in is ture, then turn #Q on and off by preset times.

   #r := SEL(G := #udt.Q,
             IN0 := #udt.time_between,
             IN1 := #udt.time_active);
   #t := "real2time_format"(in := #r, format := #udt.time_format);
   PRESET_TIMER(PT := #t, TIMER := #"timer");
   #"timer".TON(IN := #in, PT := #t, Q => #"b");

   IF NOT #in THEN
       #udt.Q := false;
       #N := 0;
   ELSIF #udt.force_off THEN
       #udt.Q := false;
   ELSIF #udt.force_on THEN
       #udt.Q := true;
   ELSIF #"b" THEN
       #udt.Q := NOT #udt.Q; // Toggle.
       #N += BOOL_TO_UINT(#udt.Q);
   END_IF;

   IF #udt.force_off OR #udt.force_on OR #"b" THEN
       RESET_TIMER(#"timer");
       #udt.force_on := false;
       #udt.force_off := false;
   END_IF;

   #RT := #"timer".PT - #"timer".ET; // Remaining time
   #udt.RT := "time2real_format"(in := #RT, format := #udt.time_format);

   #Q := #udt.Q;
END_FUNCTION_BLOCK

// folder: Library/Timers/hmi timer

FUNCTION_BLOCK "timerHmi"   // FB1, SCL
{ S7_Optimized_Access := 'TRUE' }
VERSION : 0.1
   VAR_INPUT
      in : Bool;   // Activate timer
      pt : Time;   // Added to internal "pt"
      TP : Bool;   // Puls timer
      TON : Bool;   // Timer-ON delay
      TOF : Bool;   // Timer-OFF delay
      TONR : Bool;   // Timer-ON retentiv.
   END_VAR
   VAR_OUTPUT
      Q : Bool;
      Error : Bool;   // More then one mode is active.
      RT : Time;
   END_VAR
   VAR_IN_OUT
      udt : "timerUdt";
   END_VAR
   VAR
      "timer" : IEC_TIMER;
   END_VAR
   VAR_TEMP
      p : Time;
   END_VAR
   VAR CONSTANT
      SECOUNDS : SInt;
   END_VAR
BEGIN
   // PT-max: 24 days, 20 hours, 31 min, 23 sec and 647 ms.
   // Format: 1=ms, 2=sec, 3=min, 4=h, 5=day

   // NOTE: #pt is add tho the interal preset time. (#tUdt.pt)
   #p := #pt + "real2time_format"(in := #udt.pt, format := #udt.format);

   #Error := 1 < // More then one mode is active?
   BOOL_TO_SINT(#TON) + BOOL_TO_SINT(#TOF) +
   BOOL_TO_SINT(#TP) + BOOL_TO_SINT(#TONR);

   IF #udt.format = 0 OR #Error THEN // Off
       RESET_TIMER(#"timer");
   ELSE
       // If pt is change while the timer has allread started then it will be
       // updated with the new preset time
       PRESET_TIMER(PT := #p, TIMER := #"timer");

       IF #TON THEN // Timer-ON delay
           #"timer".TON(IN := #in, PT := #p);
       ELSIF #TOF THEN // Timer-OFF delay
           #"timer".TOF(IN := #in, PT := #p);
       ELSIF #TP THEN // Puls timer
           #"timer".TP(IN := #in, PT := #p);
       ELSIF #TONR THEN // Timer-ON retentiv.
           #"timer".TONR(IN := #in, PT := #p);
       END_IF;
   END_IF;
   #Q := #"timer".Q;

   #RT := #p - #"timer".ET; // Remaining time.
   #udt.RT := "time2real_format"(in := #RT, format := #udt.format);
END_FUNCTION_BLOCK

// folder: Library/Valves

FUNCTION_BLOCK "_example_motorValve"   // FB12, SCL
{ S7_Optimized_Access := 'TRUE' }
VERSION : 0.1
   VAR_INPUT
      ai_valve1Pos : Int;
      di_valve1FullyOpen : Bool;
      di_valve1FullyClosed : Bool;
   END_VAR
   VAR_OUTPUT
      do_valve1Open : Bool;
      do_valve1Close : Bool;
   END_VAR
   VAR_IN_OUT
      ioGlobal : "ioGlobal_FB";
   END_VAR
   VAR
      valve1 : "motorValve";
      valve2 : "motorValve";
      motorValveSimulation_1 : "motorValveSimulation";
      motorValveSimulation_2 : "motorValveSimulation";
      speed : Real := 1.0;
   END_VAR
BEGIN

   // Valve 1 - (The linking block isn't required)
   "ioGlobalMotorValveLinking"(ioGlobal := #ioGlobal, valve := #valve1);
   #valve1
   (
    iFeedbackPosition := "analogInSimple"(mn := 0, in := #ai_valve1Pos, mx := 100),
    iFeddbackPosError := "analogInError"(#ai_valve1Pos),
    iFeedbackFullyOpen := #di_valve1FullyOpen,
    iFeedbackFullyClosed := #di_valve1FullyClosed,
    qOpen => #do_valve1Open,
    qClose => #do_valve1Close
   );

   // Vavle 2
   "ioGlobalMotorValveLinking"(ioGlobal := #ioGlobal, valve := #valve2);
   #valve2();

   // ---------------------------------
   // Simulation

   // IO-mapping for the valves most be commented-out, to make simulation work.
   #motorValveSimulation_1(speed := #speed, io := #valve1.hmi.io);
   #motorValveSimulation_2(speed := #speed, io := #valve2.hmi.io);
END_FUNCTION_BLOCK

// folder: Library/Valves/Blocks and UDT's

FUNCTION_BLOCK "motorValveCtrl"   // FB9, SCL
{ S7_Optimized_Access := 'TRUE' }
VERSION : 0.1
   VAR_INPUT
      iSP : Real;   // 0-100 %,
      iFailSafe : Bool;   // Open or close the valve entirly, set inside conf.
      iInterlook : Bool;   // Stop movement, valve will continue when input is set back false.
      iStop : Bool;   // Stop movement, also after var. is back false.
      iJogOpen : Bool;   // Move the valve towards open when true, has priority over SP.
      iJogClose : Bool;   // Move the valve towards close when true, has priority over SP.
      iMan : Bool := true;   // 0=auto
      iReset : Bool;   // Reset timeout.
      iRegMode : Bool;   // Most be set true, if valve is controlled by a PID.
      iExternalError : Bool;
   END_VAR
   VAR_OUTPUT
      qTimeout : Bool;   // (quick and long timeout)
   END_VAR
   VAR_IN_OUT
      conf : "motorValveConfUdt";   // Configuration parameters
      io : "motorValveIoUdt";   // Fyzical in- and outputs.
   END_VAR
   VAR
      statIn : Struct
         fullyOpen : Bool;
         fullyClosed : Bool;
      END_STRUCT;
      out : Struct
         qucikTimeout : Bool;
         longTimeout : Bool;
      END_STRUCT;
      action : SInt;   // 1=open, 2=close
      action2 : SInt;
      old : Struct
         action : SInt;
         action2 : SInt;
         SP : Real;
      END_STRUCT;
      RTRIG_iFailSafe : R_TRIG;
      RTIRG_iReset : R_TRIG;
      RTIRG_jog : R_TRIG;
      RTIRG_auto : R_TRIG;
      RTRIG_iInterlook_released : R_TRIG;
      RTRIG_iFailSafe_released : R_TRIG;
      RTRIG_jogOpen_released : R_TRIG;
      RTRIG_jogClose_released : R_TRIG;
      TP_toggleOut : IEC_TIMER;
      TON_gentle : IEC_TIMER;
      TON_regModeWait : IEC_TIMER;
      TONR_timeout : IEC_TIMER;
      TONR_quckTimeoutInterval : IEC_TIMER;
      quickTimeoutLastPos : Real;
      gentleAction : Bool;
      gentleMode : Bool;
      bothSensors : Struct
         open : Bool;
         closed : Bool;
      END_STRUCT;
   END_VAR
   VAR_TEMP
      pre : Real;
      pause : Time;
      g : Bool;
   END_VAR
   VAR CONSTANT
      NO_ACTION : SInt := 0;
      OPEN : SInt := 1;
      CLOSE : SInt := 2;
   END_VAR
BEGIN
   // Valve with analog feedback.

   // v0.1.0

   // This block doesn't include any functionality for auto-man, the reason for this 
   // is because this functionality varies from project to project.

   REGION End-pos-switches
       // Use the position signal instead of the end-limit-switches to 
       // determined if the valve is fully open or fully closed.
       // Usefull if the valve dosen't have end-limit-switches or a
       // switch dosen't work and temperary quick fix is needed.
       #statIn.fullyOpen := SEL(G := #conf.simFullyOpenWithPos,
                                IN0 := #io.in.fullyOpen,
                                IN1 := #io.in.pos > #conf.fullyOpenPosLim
                                AND NOT #io.in.posError);
       #statIn.fullyClosed := SEL(G := #conf.simFullyClosedWithPos,
                                  IN0 := #io.in.fullyClosed,
                                  IN1 := #io.in.pos < #conf.fullyClosedPosLim
                                  AND NOT #io.in.posError);

       // Two signals, both the posistion sensor and end limit sensor. If above 
       // feature is disabled.
       #bothSensors.open := (#io.in.fullyOpen OR #conf.simFullyOpenWithPos)
       (* *)AND #io.in.pos > #conf.fullyOpenPosLim AND NOT #io.in.posError;
       #bothSensors.closed := (#io.in.fullyClosed OR #conf.simFullyClosedWithPos)
       (* *)AND #io.in.pos < #conf.fullyClosedPosLim AND NOT #io.in.posError;
   END_REGION

